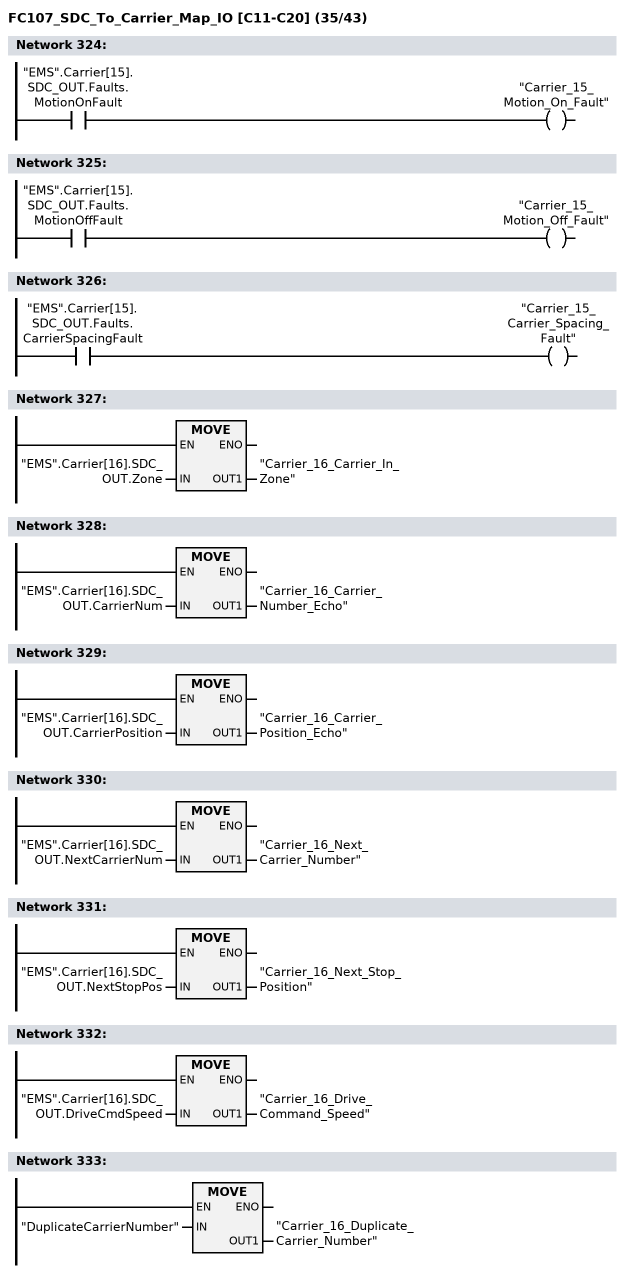
   RUNG wire#powerrail
      Contact( "EMS".Carrier[15].SDC_OUT.Faults.MotionOnFault )
      Coil( "Carrier_15_Motion_On_Fault" )
   END_RUNG
   // the same network as SCL:
   "Carrier_15_Motion_On_Fault" := "EMS".Carrier[15].SDC_OUT.Faults.MotionOnFault;
END_REGION

REGION Network 325
   RUNG wire#powerrail
      Contact( "EMS".Carrier[15].SDC_OUT.Faults.MotionOffFault )
      Coil( "Carrier_15_Motion_Off_Fault" )
   END_RUNG
   // the same network as SCL:
   "Carrier_15_Motion_Off_Fault" := "EMS".Carrier[15].SDC_OUT.Faults.MotionOffFault;
END_REGION

REGION Network 326
   RUNG wire#powerrail
      Contact( "EMS".Carrier[15].SDC_OUT.Faults.CarrierSpacingFault )
      Coil( "Carrier_15_Carrier_Spacing_Fault" )
   END_RUNG
   // the same network as SCL:
   "Carrier_15_Carrier_Spacing_Fault" := "EMS".Carrier[15].SDC_OUT.Faults.CarrierSpacingFault;
END_REGION

REGION Network 327
   RUNG wire#powerrail
      Move(in := "EMS".Carrier[16].SDC_OUT.Zone, out1 => "Carrier_16_Carrier_In_Zone")
   END_RUNG
   // the same network as SCL:
   "Carrier_16_Carrier_In_Zone" := "EMS".Carrier[16].SDC_OUT.Zone;
END_REGION

REGION Network 328
   RUNG wire#powerrail
      Move(in := "EMS".Carrier[16].SDC_OUT.CarrierNum, out1 => "Carrier_16_Carrier_Number_Echo")
   END_RUNG
   // the same network as SCL:
   "Carrier_16_Carrier_Number_Echo" := "EMS".Carrier[16].SDC_OUT.CarrierNum;
END_REGION

REGION Network 329
   RUNG wire#powerrail
      Move(in := "EMS".Carrier[16].SDC_OUT.CarrierPosition, out1 => "Carrier_16_Carrier_Position_Echo")
   END_RUNG
   // the same network as SCL:
   "Carrier_16_Carrier_Position_Echo" := "EMS".Carrier[16].SDC_OUT.CarrierPosition;
END_REGION

REGION Network 330
   RUNG wire#powerrail
      Move(in := "EMS".Carrier[16].SDC_OUT.NextCarrierNum, out1 => "Carrier_16_Next_Carrier_Number")
   END_RUNG
   // the same network as SCL:
   "Carrier_16_Next_Carrier_Number" := "EMS".Carrier[16].SDC_OUT.NextCarrierNum;
END_REGION

REGION Network 331
   RUNG wire#powerrail
      Move(in := "EMS".Carrier[16].SDC_OUT.NextStopPos, out1 => "Carrier_16_Next_Stop_Position")
   END_RUNG
   // the same network as SCL:
   "Carrier_16_Next_Stop_Position" := "EMS".Carrier[16].SDC_OUT.NextStopPos;
END_REGION

REGION Network 332
   RUNG wire#powerrail
      Move(in := "EMS".Carrier[16].SDC_OUT.DriveCmdSpeed, out1 => "Carrier_16_Drive_Command_Speed")
   END_RUNG
   // the same network as SCL:
   "Carrier_16_Drive_Command_Speed" := "EMS".Carrier[16].SDC_OUT.DriveCmdSpeed;
END_REGION

REGION Network 333
   RUNG wire#powerrail
      Move(in := "DuplicateCarrierNumber", out1 => "Carrier_16_Duplicate_Carrier_Number")
   END_RUNG
   // the same network as SCL:
   "Carrier_16_Duplicate_Carrier_Number" := "DuplicateCarrierNumber";
END_REGION

REGION Network 334
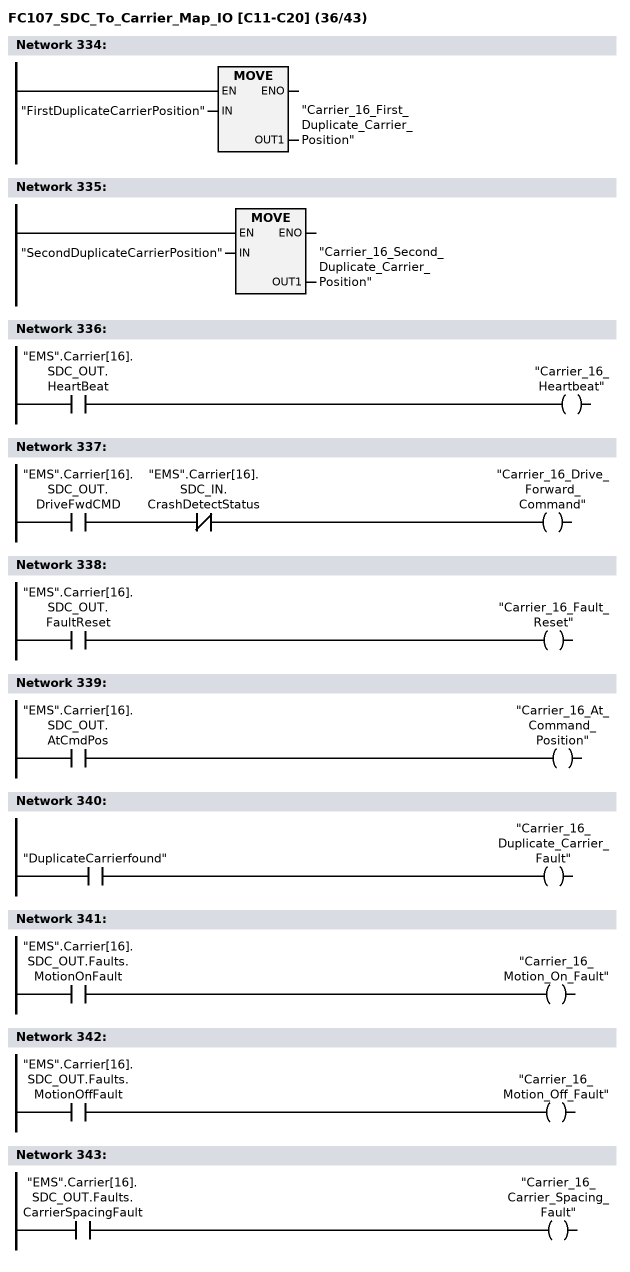
   RUNG wire#powerrail
      Move(in := "FirstDuplicateCarrierPosition", out1 => "Carrier_16_First_Duplicate_Carrier_Position")
   END_RUNG
   // the same network as SCL:
   "Carrier_16_First_Duplicate_Carrier_Position" := "FirstDuplicateCarrierPosition";
END_REGION

REGION Network 335
   RUNG wire#powerrail
      Move(in := "SecondDuplicateCarrierPosition", out1 => "Carrier_16_Second_Duplicate_Carrier_Position")
   END_RUNG
   // the same network as SCL:
   "Carrier_16_Second_Duplicate_Carrier_Position" := "SecondDuplicateCarrierPosition";
END_REGION

REGION Network 336
   RUNG wire#powerrail
      Contact( "EMS".Carrier[16].SDC_OUT.HeartBeat )
      Coil( "Carrier_16_Heartbeat" )
   END_RUNG
   // the same network as SCL:
   "Carrier_16_Heartbeat" := "EMS".Carrier[16].SDC_OUT.HeartBeat;
END_REGION

REGION Network 337
   RUNG wire#powerrail
      Contact( "EMS".Carrier[16].SDC_OUT.DriveFwdCMD )
      I_Contact( "EMS".Carrier[16].SDC_IN.CrashDetectStatus )
      Coil( "Carrier_16_Drive_Forward_Command" )
   END_RUNG
   // the same network as SCL:
   "Carrier_16_Drive_Forward_Command" := "EMS".Carrier[16].SDC_OUT.DriveFwdCMD AND NOT "EMS".Carrier[16].SDC_IN.CrashDetectStatus;
END_REGION

REGION Network 338
   RUNG wire#powerrail
      Contact( "EMS".Carrier[16].SDC_OUT.FaultReset )
      Coil( "Carrier_16_Fault_Reset" )
   END_RUNG
   // the same network as SCL:
   "Carrier_16_Fault_Reset" := "EMS".Carrier[16].SDC_OUT.FaultReset;
END_REGION

REGION Network 339
   RUNG wire#powerrail
      Contact( "EMS".Carrier[16].SDC_OUT.AtCmdPos )
      Coil( "Carrier_16_At_Command_Position" )
   END_RUNG
   // the same network as SCL:
   "Carrier_16_At_Command_Position" := "EMS".Carrier[16].SDC_OUT.AtCmdPos;
END_REGION

REGION Network 340
   RUNG wire#powerrail
      Contact( "DuplicateCarrierfound" )
      Coil( "Carrier_16_Duplicate_Carrier_Fault" )
   END_RUNG
   // the same network as SCL:
   "Carrier_16_Duplicate_Carrier_Fault" := "DuplicateCarrierfound";
END_REGION

REGION Network 341
   RUNG wire#powerrail
      Contact( "EMS".Carrier[16].SDC_OUT.Faults.MotionOnFault )
      Coil( "Carrier_16_Motion_On_Fault" )
   END_RUNG
   // the same network as SCL:
   "Carrier_16_Motion_On_Fault" := "EMS".Carrier[16].SDC_OUT.Faults.MotionOnFault;
END_REGION

REGION Network 342
   RUNG wire#powerrail
      Contact( "EMS".Carrier[16].SDC_OUT.Faults.MotionOffFault )
      Coil( "Carrier_16_Motion_Off_Fault" )
   END_RUNG
   // the same network as SCL:
   "Carrier_16_Motion_Off_Fault" := "EMS".Carrier[16].SDC_OUT.Faults.MotionOffFault;
END_REGION

REGION Network 343
   RUNG wire#powerrail
      Contact( "EMS".Carrier[16].SDC_OUT.Faults.CarrierSpacingFault )
      Coil( "Carrier_16_Carrier_Spacing_Fault" )
   END_RUNG
   // the same network as SCL:
   "Carrier_16_Carrier_Spacing_Fault" := "EMS".Carrier[16].SDC_OUT.Faults.CarrierSpacingFault;
END_REGION

REGION Network 344
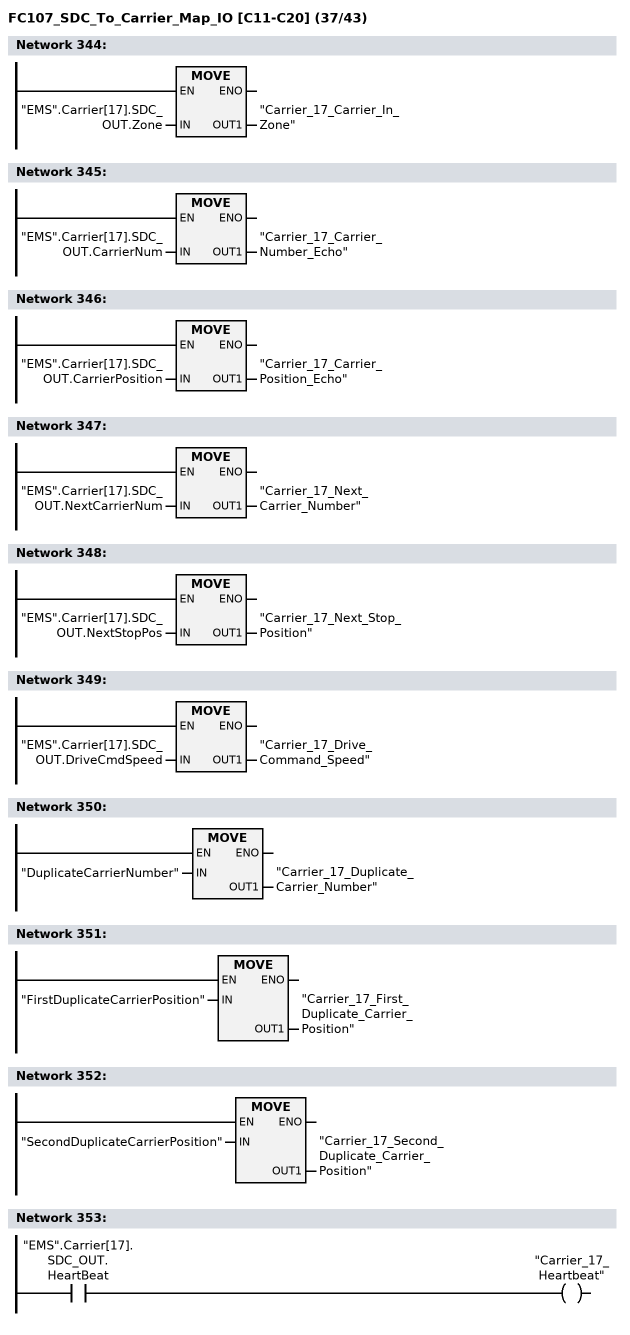
   RUNG wire#powerrail
      Move(in := "EMS".Carrier[17].SDC_OUT.Zone, out1 => "Carrier_17_Carrier_In_Zone")
   END_RUNG
   // the same network as SCL:
   "Carrier_17_Carrier_In_Zone" := "EMS".Carrier[17].SDC_OUT.Zone;
END_REGION

REGION Network 345
   RUNG wire#powerrail
      Move(in := "EMS".Carrier[17].SDC_OUT.CarrierNum, out1 => "Carrier_17_Carrier_Number_Echo")
   END_RUNG
   // the same network as SCL:
   "Carrier_17_Carrier_Number_Echo" := "EMS".Carrier[17].SDC_OUT.CarrierNum;
END_REGION

REGION Network 346
   RUNG wire#powerrail
      Move(in := "EMS".Carrier[17].SDC_OUT.CarrierPosition, out1 => "Carrier_17_Carrier_Position_Echo")
   END_RUNG
   // the same network as SCL:
   "Carrier_17_Carrier_Position_Echo" := "EMS".Carrier[17].SDC_OUT.CarrierPosition;
END_REGION

REGION Network 347
   RUNG wire#powerrail
      Move(in := "EMS".Carrier[17].SDC_OUT.NextCarrierNum, out1 => "Carrier_17_Next_Carrier_Number")
   END_RUNG
   // the same network as SCL:
   "Carrier_17_Next_Carrier_Number" := "EMS".Carrier[17].SDC_OUT.NextCarrierNum;
END_REGION

REGION Network 348
   RUNG wire#powerrail
      Move(in := "EMS".Carrier[17].SDC_OUT.NextStopPos, out1 => "Carrier_17_Next_Stop_Position")
   END_RUNG
   // the same network as SCL:
   "Carrier_17_Next_Stop_Position" := "EMS".Carrier[17].SDC_OUT.NextStopPos;
END_REGION

REGION Network 349
   RUNG wire#powerrail
      Move(in := "EMS".Carrier[17].SDC_OUT.DriveCmdSpeed, out1 => "Carrier_17_Drive_Command_Speed")
   END_RUNG
   // the same network as SCL:
   "Carrier_17_Drive_Command_Speed" := "EMS".Carrier[17].SDC_OUT.DriveCmdSpeed;
END_REGION

REGION Network 350
   RUNG wire#powerrail
      Move(in := "DuplicateCarrierNumber", out1 => "Carrier_17_Duplicate_Carrier_Number")
   END_RUNG
   // the same network as SCL:
   "Carrier_17_Duplicate_Carrier_Number" := "DuplicateCarrierNumber";
END_REGION

REGION Network 351
   RUNG wire#powerrail
      Move(in := "FirstDuplicateCarrierPosition", out1 => "Carrier_17_First_Duplicate_Carrier_Position")
   END_RUNG
   // the same network as SCL:
   "Carrier_17_First_Duplicate_Carrier_Position" := "FirstDuplicateCarrierPosition";
END_REGION

REGION Network 352
   RUNG wire#powerrail
      Move(in := "SecondDuplicateCarrierPosition", out1 => "Carrier_17_Second_Duplicate_Carrier_Position")
   END_RUNG
   // the same network as SCL:
   "Carrier_17_Second_Duplicate_Carrier_Position" := "SecondDuplicateCarrierPosition";
END_REGION

REGION Network 353
   RUNG wire#powerrail
      Contact( "EMS".Carrier[17].SDC_OUT.HeartBeat )
      Coil( "Carrier_17_Heartbeat" )
   END_RUNG
   // the same network as SCL:
   "Carrier_17_Heartbeat" := "EMS".Carrier[17].SDC_OUT.HeartBeat;
END_REGION

REGION Network 354
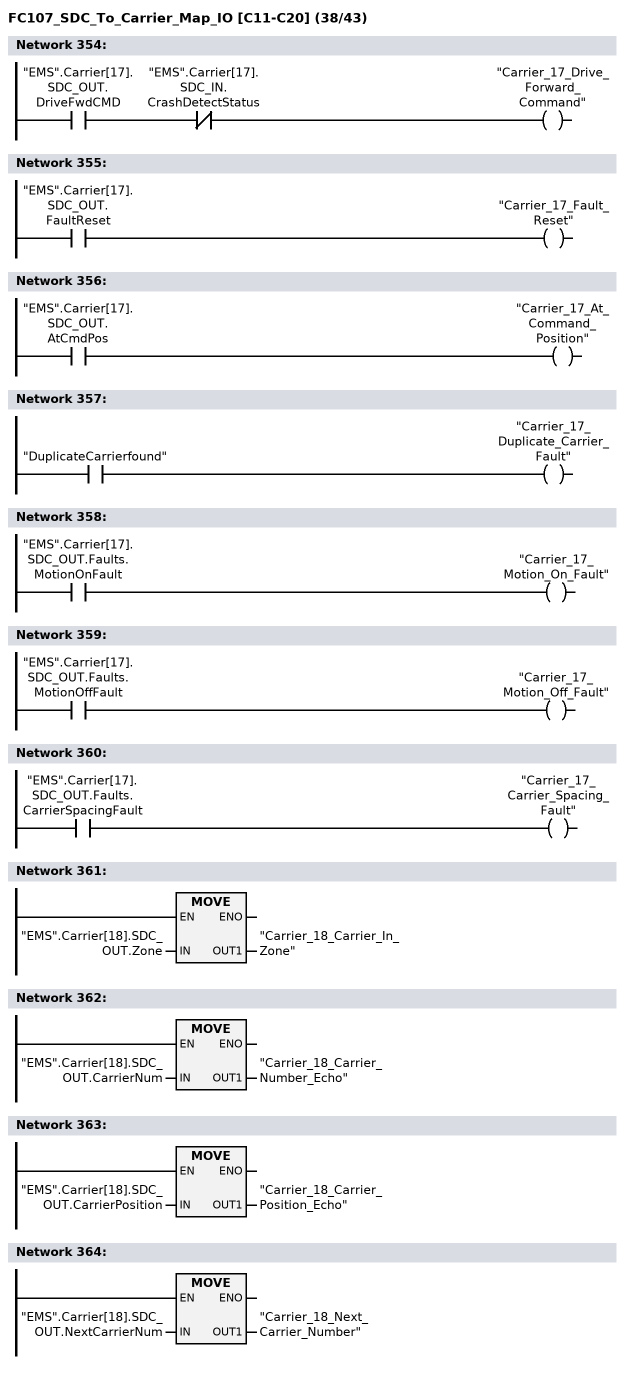
   RUNG wire#powerrail
      Contact( "EMS".Carrier[17].SDC_OUT.DriveFwdCMD )
      I_Contact( "EMS".Carrier[17].SDC_IN.CrashDetectStatus )
      Coil( "Carrier_17_Drive_Forward_Command" )
   END_RUNG
   // the same network as SCL:
   "Carrier_17_Drive_Forward_Command" := "EMS".Carrier[17].SDC_OUT.DriveFwdCMD AND NOT "EMS".Carrier[17].SDC_IN.CrashDetectStatus;
END_REGION

REGION Network 355
   RUNG wire#powerrail
      Contact( "EMS".Carrier[17].SDC_OUT.FaultReset )
      Coil( "Carrier_17_Fault_Reset" )
   END_RUNG
   // the same network as SCL:
   "Carrier_17_Fault_Reset" := "EMS".Carrier[17].SDC_OUT.FaultReset;
END_REGION

REGION Network 356
   RUNG wire#powerrail
      Contact( "EMS".Carrier[17].SDC_OUT.AtCmdPos )
      Coil( "Carrier_17_At_Command_Position" )
   END_RUNG
   // the same network as SCL:
   "Carrier_17_At_Command_Position" := "EMS".Carrier[17].SDC_OUT.AtCmdPos;
END_REGION

REGION Network 357
   RUNG wire#powerrail
      Contact( "DuplicateCarrierfound" )
      Coil( "Carrier_17_Duplicate_Carrier_Fault" )
   END_RUNG
   // the same network as SCL:
   "Carrier_17_Duplicate_Carrier_Fault" := "DuplicateCarrierfound";
END_REGION

REGION Network 358
   RUNG wire#powerrail
      Contact( "EMS".Carrier[17].SDC_OUT.Faults.MotionOnFault )
      Coil( "Carrier_17_Motion_On_Fault" )
   END_RUNG
   // the same network as SCL:
   "Carrier_17_Motion_On_Fault" := "EMS".Carrier[17].SDC_OUT.Faults.MotionOnFault;
END_REGION

REGION Network 359
   RUNG wire#powerrail
      Contact( "EMS".Carrier[17].SDC_OUT.Faults.MotionOffFault )
      Coil( "Carrier_17_Motion_Off_Fault" )
   END_RUNG
   // the same network as SCL:
   "Carrier_17_Motion_Off_Fault" := "EMS".Carrier[17].SDC_OUT.Faults.MotionOffFault;
END_REGION

REGION Network 360
   RUNG wire#powerrail
      Contact( "EMS".Carrier[17].SDC_OUT.Faults.CarrierSpacingFault )
      Coil( "Carrier_17_Carrier_Spacing_Fault" )
   END_RUNG
   // the same network as SCL:
   "Carrier_17_Carrier_Spacing_Fault" := "EMS".Carrier[17].SDC_OUT.Faults.CarrierSpacingFault;
END_REGION

REGION Network 361
   RUNG wire#powerrail
      Move(in := "EMS".Carrier[18].SDC_OUT.Zone, out1 => "Carrier_18_Carrier_In_Zone")
   END_RUNG
   // the same network as SCL:
   "Carrier_18_Carrier_In_Zone" := "EMS".Carrier[18].SDC_OUT.Zone;
END_REGION

REGION Network 362
   RUNG wire#powerrail
      Move(in := "EMS".Carrier[18].SDC_OUT.CarrierNum, out1 => "Carrier_18_Carrier_Number_Echo")
   END_RUNG
   // the same network as SCL:
   "Carrier_18_Carrier_Number_Echo" := "EMS".Carrier[18].SDC_OUT.CarrierNum;
END_REGION

REGION Network 363
   RUNG wire#powerrail
      Move(in := "EMS".Carrier[18].SDC_OUT.CarrierPosition, out1 => "Carrier_18_Carrier_Position_Echo")
   END_RUNG
   // the same network as SCL:
   "Carrier_18_Carrier_Position_Echo" := "EMS".Carrier[18].SDC_OUT.CarrierPosition;
END_REGION

REGION Network 364
   RUNG wire#powerrail
      Move(in := "EMS".Carrier[18].SDC_OUT.NextCarrierNum, out1 => "Carrier_18_Next_Carrier_Number")
   END_RUNG
   // the same network as SCL:
   "Carrier_18_Next_Carrier_Number" := "EMS".Carrier[18].SDC_OUT.NextCarrierNum;
END_REGION

REGION Network 365
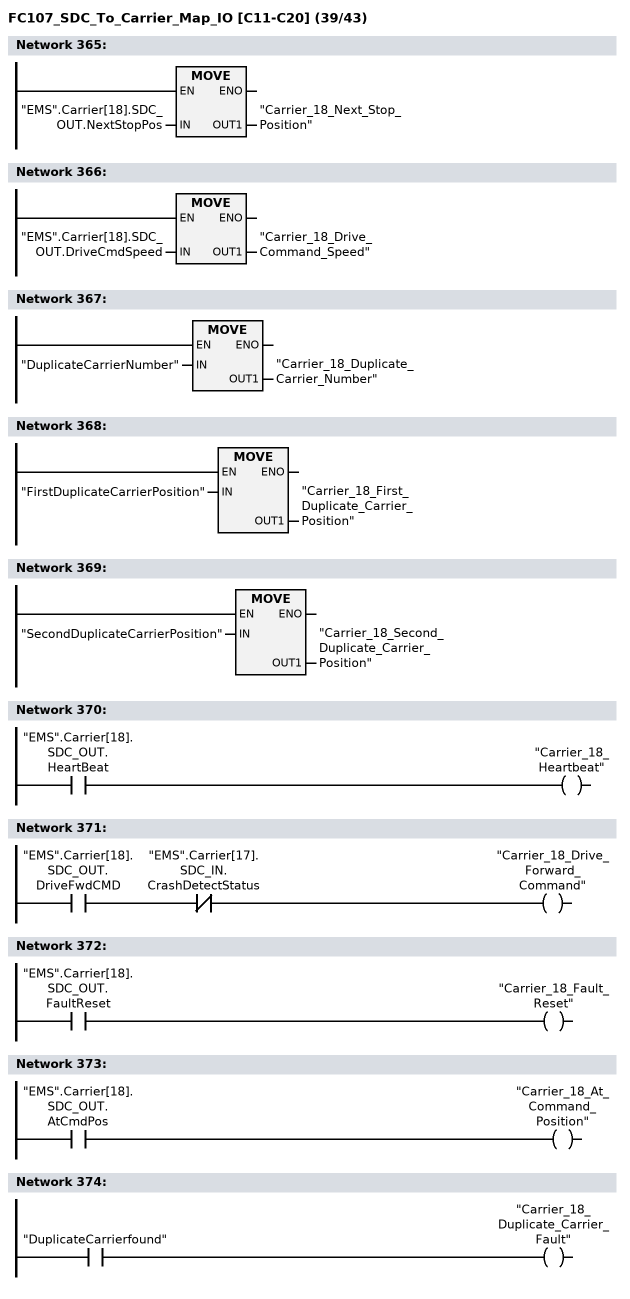
   RUNG wire#powerrail
      Move(in := "EMS".Carrier[18].SDC_OUT.NextStopPos, out1 => "Carrier_18_Next_Stop_Position")
   END_RUNG
   // the same network as SCL:
   "Carrier_18_Next_Stop_Position" := "EMS".Carrier[18].SDC_OUT.NextStopPos;
END_REGION

REGION Network 366
   RUNG wire#powerrail
      Move(in := "EMS".Carrier[18].SDC_OUT.DriveCmdSpeed, out1 => "Carrier_18_Drive_Command_Speed")
   END_RUNG
   // the same network as SCL:
   "Carrier_18_Drive_Command_Speed" := "EMS".Carrier[18].SDC_OUT.DriveCmdSpeed;
END_REGION

REGION Network 367
   RUNG wire#powerrail
      Move(in := "DuplicateCarrierNumber", out1 => "Carrier_18_Duplicate_Carrier_Number")
   END_RUNG
   // the same network as SCL:
   "Carrier_18_Duplicate_Carrier_Number" := "DuplicateCarrierNumber";
END_REGION

REGION Network 368
   RUNG wire#powerrail
      Move(in := "FirstDuplicateCarrierPosition", out1 => "Carrier_18_First_Duplicate_Carrier_Position")
   END_RUNG
   // the same network as SCL:
   "Carrier_18_First_Duplicate_Carrier_Position" := "FirstDuplicateCarrierPosition";
END_REGION

REGION Network 369
   RUNG wire#powerrail
      Move(in := "SecondDuplicateCarrierPosition", out1 => "Carrier_18_Second_Duplicate_Carrier_Position")
   END_RUNG
   // the same network as SCL:
   "Carrier_18_Second_Duplicate_Carrier_Position" := "SecondDuplicateCarrierPosition";
END_REGION

REGION Network 370
   RUNG wire#powerrail
      Contact( "EMS".Carrier[18].SDC_OUT.HeartBeat )
      Coil( "Carrier_18_Heartbeat" )
   END_RUNG
   // the same network as SCL:
   "Carrier_18_Heartbeat" := "EMS".Carrier[18].SDC_OUT.HeartBeat;
END_REGION

REGION Network 371
   RUNG wire#powerrail
      Contact( "EMS".Carrier[18].SDC_OUT.DriveFwdCMD )
      I_Contact( "EMS".Carrier[17].SDC_IN.CrashDetectStatus )
      Coil( "Carrier_18_Drive_Forward_Command" )
   END_RUNG
   // the same network as SCL:
   "Carrier_18_Drive_Forward_Command" := "EMS".Carrier[18].SDC_OUT.DriveFwdCMD AND NOT "EMS".Carrier[17].SDC_IN.CrashDetectStatus;
END_REGION

REGION Network 372
   RUNG wire#powerrail
      Contact( "EMS".Carrier[18].SDC_OUT.FaultReset )
      Coil( "Carrier_18_Fault_Reset" )
   END_RUNG
   // the same network as SCL:
   "Carrier_18_Fault_Reset" := "EMS".Carrier[18].SDC_OUT.FaultReset;
END_REGION

REGION Network 373
   RUNG wire#powerrail
      Contact( "EMS".Carrier[18].SDC_OUT.AtCmdPos )
      Coil( "Carrier_18_At_Command_Position" )
   END_RUNG
   // the same network as SCL:
   "Carrier_18_At_Command_Position" := "EMS".Carrier[18].SDC_OUT.AtCmdPos;
END_REGION

REGION Network 374
   RUNG wire#powerrail
      Contact( "DuplicateCarrierfound" )
      Coil( "Carrier_18_Duplicate_Carrier_Fault" )
   END_RUNG
   // the same network as SCL:
   "Carrier_18_Duplicate_Carrier_Fault" := "DuplicateCarrierfound";
END_REGION

REGION Network 375
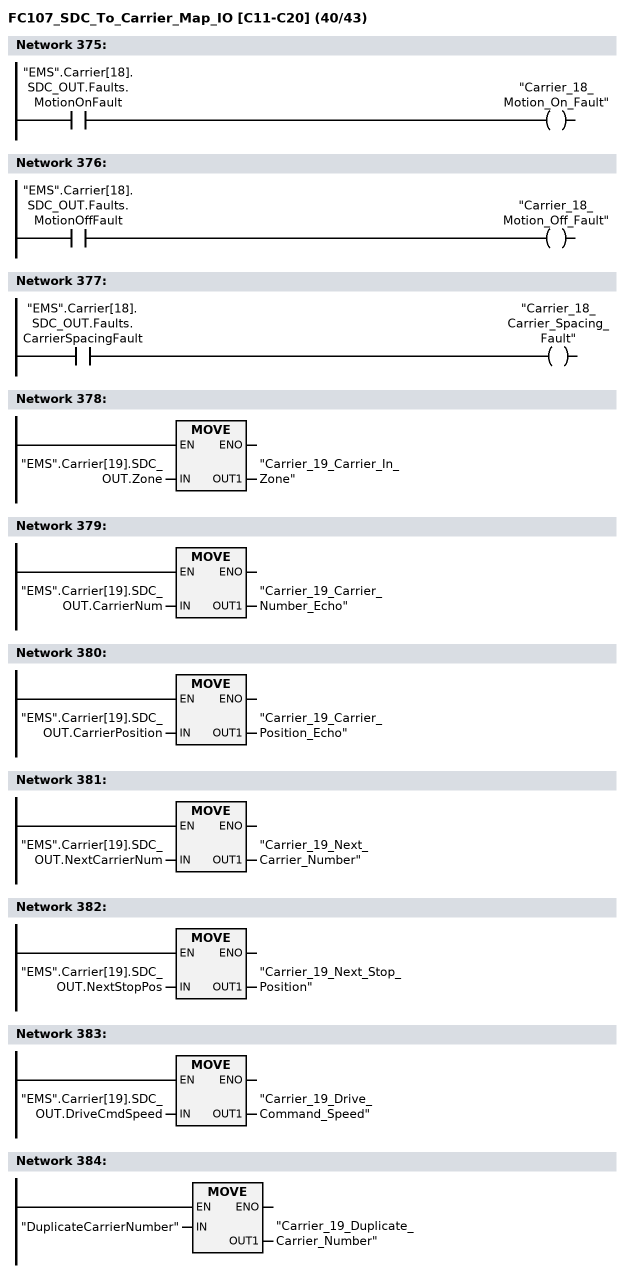
   RUNG wire#powerrail
      Contact( "EMS".Carrier[18].SDC_OUT.Faults.MotionOnFault )
      Coil( "Carrier_18_Motion_On_Fault" )
   END_RUNG
   // the same network as SCL:
   "Carrier_18_Motion_On_Fault" := "EMS".Carrier[18].SDC_OUT.Faults.MotionOnFault;
END_REGION

REGION Network 376
   RUNG wire#powerrail
      Contact( "EMS".Carrier[18].SDC_OUT.Faults.MotionOffFault )
      Coil( "Carrier_18_Motion_Off_Fault" )
   END_RUNG
   // the same network as SCL:
   "Carrier_18_Motion_Off_Fault" := "EMS".Carrier[18].SDC_OUT.Faults.MotionOffFault;
END_REGION

REGION Network 377
   RUNG wire#powerrail
      Contact( "EMS".Carrier[18].SDC_OUT.Faults.CarrierSpacingFault )
      Coil( "Carrier_18_Carrier_Spacing_Fault" )
   END_RUNG
   // the same network as SCL:
   "Carrier_18_Carrier_Spacing_Fault" := "EMS".Carrier[18].SDC_OUT.Faults.CarrierSpacingFault;
END_REGION

REGION Network 378
   RUNG wire#powerrail
      Move(in := "EMS".Carrier[19].SDC_OUT.Zone, out1 => "Carrier_19_Carrier_In_Zone")
   END_RUNG
   // the same network as SCL:
   "Carrier_19_Carrier_In_Zone" := "EMS".Carrier[19].SDC_OUT.Zone;
END_REGION

REGION Network 379
   RUNG wire#powerrail
      Move(in := "EMS".Carrier[19].SDC_OUT.CarrierNum, out1 => "Carrier_19_Carrier_Number_Echo")
   END_RUNG
   // the same network as SCL:
   "Carrier_19_Carrier_Number_Echo" := "EMS".Carrier[19].SDC_OUT.CarrierNum;
END_REGION

REGION Network 380
   RUNG wire#powerrail
      Move(in := "EMS".Carrier[19].SDC_OUT.CarrierPosition, out1 => "Carrier_19_Carrier_Position_Echo")
   END_RUNG
   // the same network as SCL:
   "Carrier_19_Carrier_Position_Echo" := "EMS".Carrier[19].SDC_OUT.CarrierPosition;
END_REGION

REGION Network 381
   RUNG wire#powerrail
      Move(in := "EMS".Carrier[19].SDC_OUT.NextCarrierNum, out1 => "Carrier_19_Next_Carrier_Number")
   END_RUNG
   // the same network as SCL:
   "Carrier_19_Next_Carrier_Number" := "EMS".Carrier[19].SDC_OUT.NextCarrierNum;
END_REGION

REGION Network 382
   RUNG wire#powerrail
      Move(in := "EMS".Carrier[19].SDC_OUT.NextStopPos, out1 => "Carrier_19_Next_Stop_Position")
   END_RUNG
   // the same network as SCL:
   "Carrier_19_Next_Stop_Position" := "EMS".Carrier[19].SDC_OUT.NextStopPos;
END_REGION

REGION Network 383
   RUNG wire#powerrail
      Move(in := "EMS".Carrier[19].SDC_OUT.DriveCmdSpeed, out1 => "Carrier_19_Drive_Command_Speed")
   END_RUNG
   // the same network as SCL:
   "Carrier_19_Drive_Command_Speed" := "EMS".Carrier[19].SDC_OUT.DriveCmdSpeed;
END_REGION

REGION Network 384
   RUNG wire#powerrail
      Move(in := "DuplicateCarrierNumber", out1 => "Carrier_19_Duplicate_Carrier_Number")
   END_RUNG
   // the same network as SCL:
   "Carrier_19_Duplicate_Carrier_Number" := "DuplicateCarrierNumber";
END_REGION

REGION Network 385
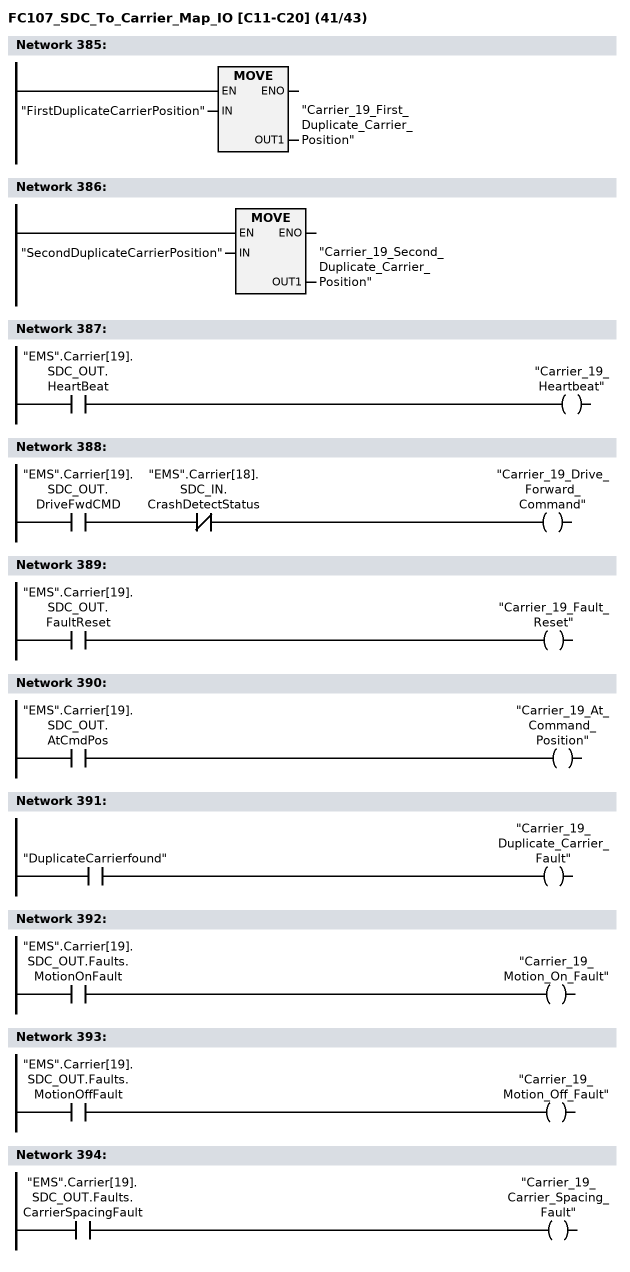
   RUNG wire#powerrail
      Move(in := "FirstDuplicateCarrierPosition", out1 => "Carrier_19_First_Duplicate_Carrier_Position")
   END_RUNG
   // the same network as SCL:
   "Carrier_19_First_Duplicate_Carrier_Position" := "FirstDuplicateCarrierPosition";
END_REGION

REGION Network 386
   RUNG wire#powerrail
      Move(in := "SecondDuplicateCarrierPosition", out1 => "Carrier_19_Second_Duplicate_Carrier_Position")
   END_RUNG
   // the same network as SCL:
   "Carrier_19_Second_Duplicate_Carrier_Position" := "SecondDuplicateCarrierPosition";
END_REGION

REGION Network 387
   RUNG wire#powerrail
      Contact( "EMS".Carrier[19].SDC_OUT.HeartBeat )
      Coil( "Carrier_19_Heartbeat" )
   END_RUNG
   // the same network as SCL:
   "Carrier_19_Heartbeat" := "EMS".Carrier[19].SDC_OUT.HeartBeat;
END_REGION

REGION Network 388
   RUNG wire#powerrail
      Contact( "EMS".Carrier[19].SDC_OUT.DriveFwdCMD )
      I_Contact( "EMS".Carrier[18].SDC_IN.CrashDetectStatus )
      Coil( "Carrier_19_Drive_Forward_Command" )
   END_RUNG
   // the same network as SCL:
   "Carrier_19_Drive_Forward_Command" := "EMS".Carrier[19].SDC_OUT.DriveFwdCMD AND NOT "EMS".Carrier[18].SDC_IN.CrashDetectStatus;
END_REGION

REGION Network 389
   RUNG wire#powerrail
      Contact( "EMS".Carrier[19].SDC_OUT.FaultReset )
      Coil( "Carrier_19_Fault_Reset" )
   END_RUNG
   // the same network as SCL:
   "Carrier_19_Fault_Reset" := "EMS".Carrier[19].SDC_OUT.FaultReset;
END_REGION

REGION Network 390
   RUNG wire#powerrail
      Contact( "EMS".Carrier[19].SDC_OUT.AtCmdPos )
      Coil( "Carrier_19_At_Command_Position" )
   END_RUNG
   // the same network as SCL:
   "Carrier_19_At_Command_Position" := "EMS".Carrier[19].SDC_OUT.AtCmdPos;
END_REGION

REGION Network 391
   RUNG wire#powerrail
      Contact( "DuplicateCarrierfound" )
      Coil( "Carrier_19_Duplicate_Carrier_Fault" )
   END_RUNG
   // the same network as SCL:
   "Carrier_19_Duplicate_Carrier_Fault" := "DuplicateCarrierfound";
END_REGION

REGION Network 392
   RUNG wire#powerrail
      Contact( "EMS".Carrier[19].SDC_OUT.Faults.MotionOnFault )
      Coil( "Carrier_19_Motion_On_Fault" )
   END_RUNG
   // the same network as SCL:
   "Carrier_19_Motion_On_Fault" := "EMS".Carrier[19].SDC_OUT.Faults.MotionOnFault;
END_REGION

REGION Network 393
   RUNG wire#powerrail
      Contact( "EMS".Carrier[19].SDC_OUT.Faults.MotionOffFault )
      Coil( "Carrier_19_Motion_Off_Fault" )
   END_RUNG
   // the same network as SCL:
   "Carrier_19_Motion_Off_Fault" := "EMS".Carrier[19].SDC_OUT.Faults.MotionOffFault;
END_REGION

REGION Network 394
   RUNG wire#powerrail
      Contact( "EMS".Carrier[19].SDC_OUT.Faults.CarrierSpacingFault )
      Coil( "Carrier_19_Carrier_Spacing_Fault" )
   END_RUNG
   // the same network as SCL:
   "Carrier_19_Carrier_Spacing_Fault" := "EMS".Carrier[19].SDC_OUT.Faults.CarrierSpacingFault;
END_REGION

REGION Network 395
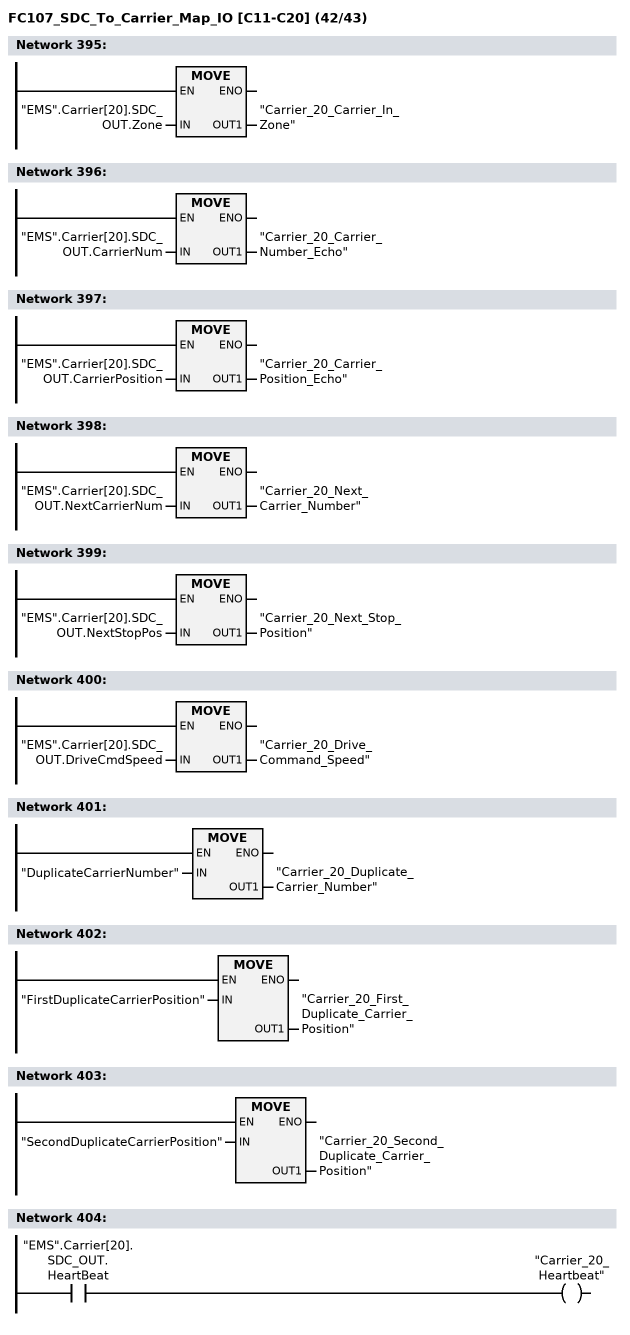
   RUNG wire#powerrail
      Move(in := "EMS".Carrier[20].SDC_OUT.Zone, out1 => "Carrier_20_Carrier_In_Zone")
   END_RUNG
   // the same network as SCL:
   "Carrier_20_Carrier_In_Zone" := "EMS".Carrier[20].SDC_OUT.Zone;
END_REGION

REGION Network 396
   RUNG wire#powerrail
      Move(in := "EMS".Carrier[20].SDC_OUT.CarrierNum, out1 => "Carrier_20_Carrier_Number_Echo")
   END_RUNG
   // the same network as SCL:
   "Carrier_20_Carrier_Number_Echo" := "EMS".Carrier[20].SDC_OUT.CarrierNum;
END_REGION

REGION Network 397
   RUNG wire#powerrail
      Move(in := "EMS".Carrier[20].SDC_OUT.CarrierPosition, out1 => "Carrier_20_Carrier_Position_Echo")
   END_RUNG
   // the same network as SCL:
   "Carrier_20_Carrier_Position_Echo" := "EMS".Carrier[20].SDC_OUT.CarrierPosition;
END_REGION

REGION Network 398
   RUNG wire#powerrail
      Move(in := "EMS".Carrier[20].SDC_OUT.NextCarrierNum, out1 => "Carrier_20_Next_Carrier_Number")
   END_RUNG
   // the same network as SCL:
   "Carrier_20_Next_Carrier_Number" := "EMS".Carrier[20].SDC_OUT.NextCarrierNum;
END_REGION

REGION Network 399
   RUNG wire#powerrail
      Move(in := "EMS".Carrier[20].SDC_OUT.NextStopPos, out1 => "Carrier_20_Next_Stop_Position")
   END_RUNG
   // the same network as SCL:
   "Carrier_20_Next_Stop_Position" := "EMS".Carrier[20].SDC_OUT.NextStopPos;
END_REGION

REGION Network 400
   RUNG wire#powerrail
      Move(in := "EMS".Carrier[20].SDC_OUT.DriveCmdSpeed, out1 => "Carrier_20_Drive_Command_Speed")
   END_RUNG
   // the same network as SCL:
   "Carrier_20_Drive_Command_Speed" := "EMS".Carrier[20].SDC_OUT.DriveCmdSpeed;
END_REGION

REGION Network 401
   RUNG wire#powerrail
      Move(in := "DuplicateCarrierNumber", out1 => "Carrier_20_Duplicate_Carrier_Number")
   END_RUNG
   // the same network as SCL:
   "Carrier_20_Duplicate_Carrier_Number" := "DuplicateCarrierNumber";
END_REGION

REGION Network 402
   RUNG wire#powerrail
      Move(in := "FirstDuplicateCarrierPosition", out1 => "Carrier_20_First_Duplicate_Carrier_Position")
   END_RUNG
   // the same network as SCL:
   "Carrier_20_First_Duplicate_Carrier_Position" := "FirstDuplicateCarrierPosition";
END_REGION

REGION Network 403
   RUNG wire#powerrail
      Move(in := "SecondDuplicateCarrierPosition", out1 => "Carrier_20_Second_Duplicate_Carrier_Position")
   END_RUNG
   // the same network as SCL:
   "Carrier_20_Second_Duplicate_Carrier_Position" := "SecondDuplicateCarrierPosition";
END_REGION

REGION Network 404
   RUNG wire#powerrail
      Contact( "EMS".Carrier[20].SDC_OUT.HeartBeat )
      Coil( "Carrier_20_Heartbeat" )
   END_RUNG
   // the same network as SCL:
   "Carrier_20_Heartbeat" := "EMS".Carrier[20].SDC_OUT.HeartBeat;
END_REGION

REGION Network 405
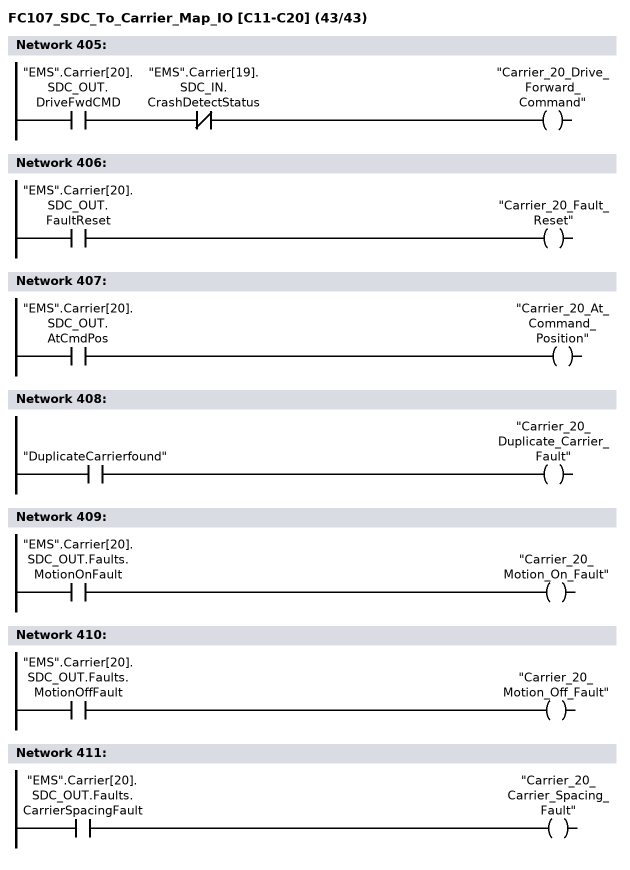
   RUNG wire#powerrail
      Contact( "EMS".Carrier[20].SDC_OUT.DriveFwdCMD )
      I_Contact( "EMS".Carrier[19].SDC_IN.CrashDetectStatus )
      Coil( "Carrier_20_Drive_Forward_Command" )
   END_RUNG
   // the same network as SCL:
   "Carrier_20_Drive_Forward_Command" := "EMS".Carrier[20].SDC_OUT.DriveFwdCMD AND NOT "EMS".Carrier[19].SDC_IN.CrashDetectStatus;
END_REGION

REGION Network 406
   RUNG wire#powerrail
      Contact( "EMS".Carrier[20].SDC_OUT.FaultReset )
      Coil( "Carrier_20_Fault_Reset" )
   END_RUNG
   // the same network as SCL:
   "Carrier_20_Fault_Reset" := "EMS".Carrier[20].SDC_OUT.FaultReset;
END_REGION

REGION Network 407
   RUNG wire#powerrail
      Contact( "EMS".Carrier[20].SDC_OUT.AtCmdPos )
      Coil( "Carrier_20_At_Command_Position" )
   END_RUNG
   // the same network as SCL:
   "Carrier_20_At_Command_Position" := "EMS".Carrier[20].SDC_OUT.AtCmdPos;
END_REGION

REGION Network 408
   RUNG wire#powerrail
      Contact( "DuplicateCarrierfound" )
      Coil( "Carrier_20_Duplicate_Carrier_Fault" )
   END_RUNG
   // the same network as SCL:
   "Carrier_20_Duplicate_Carrier_Fault" := "DuplicateCarrierfound";
END_REGION

REGION Network 409
   RUNG wire#powerrail
      Contact( "EMS".Carrier[20].SDC_OUT.Faults.MotionOnFault )
      Coil( "Carrier_20_Motion_On_Fault" )
   END_RUNG
   // the same network as SCL:
   "Carrier_20_Motion_On_Fault" := "EMS".Carrier[20].SDC_OUT.Faults.MotionOnFault;
END_REGION

REGION Network 410
   RUNG wire#powerrail
      Contact( "EMS".Carrier[20].SDC_OUT.Faults.MotionOffFault )
      Coil( "Carrier_20_Motion_Off_Fault" )
   END_RUNG
   // the same network as SCL:
   "Carrier_20_Motion_Off_Fault" := "EMS".Carrier[20].SDC_OUT.Faults.MotionOffFault;
END_REGION
